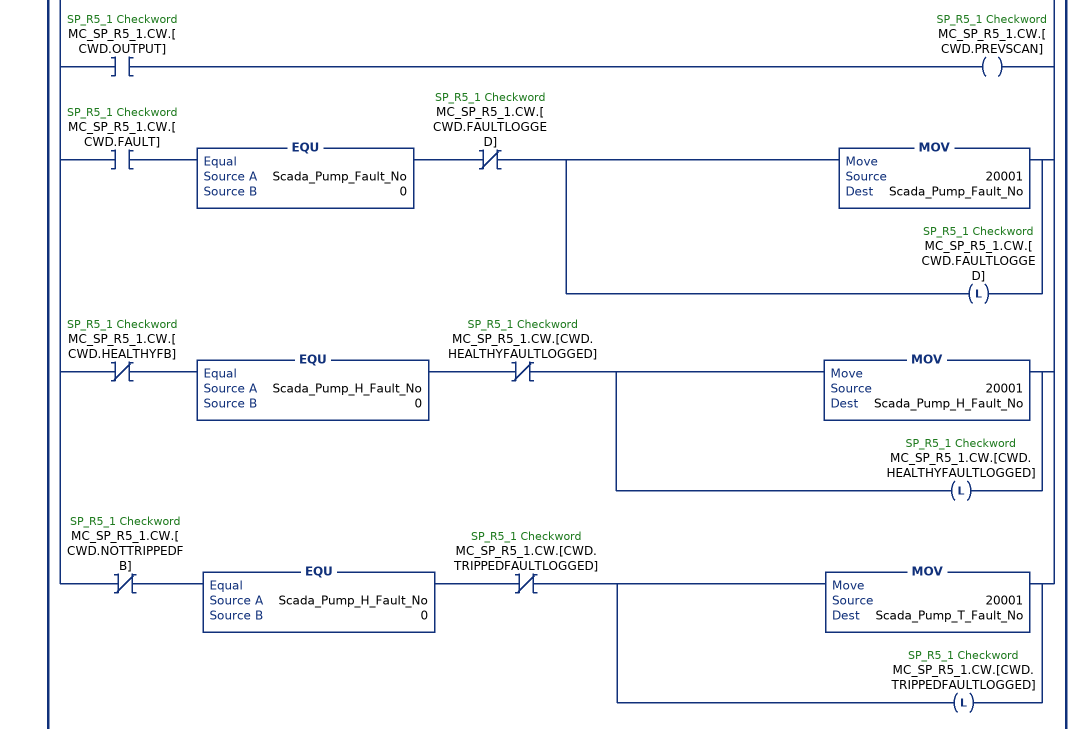
   7: [NEQ(MC_SP_R5_1.DriveBits,0) OTE(MC_SP_R5_1.CW.[CWD.AUTODRV]) ,[XIC(MC_SP_R5_1.CW.[CWD.AUTODRV]) XIO(MC_SP_R5_1.CW.[CWD.MANUAL]) ,XIC(MC_SP_R5_1.CW.[CWD.MANDRV]) XIC(MC_SP_R5_1.CW.[CWD.MANUAL]) ] OTE(MC_SP_R5_1.CW.[CWD.OUTPUT]) ,XIC(MC_SP_R5_1.CW.[CWD.OUTPUT]) OTE(MC_SP_R5_1_D) ,XIC(S:FS) [OTU(MC_SP_R5_1.CW.[CWD.MANUAL]) ,LEQ(MC_SP_R5_1.CheckTime,0) MOV(Default_Check_Time,MC_SP_R5_1.CheckTime) ] ,[[XIC(MC_SP_R5_1_R) XIO(Item_Simulation_Flag) ,XIC(Item_Simulation_Flag) [XIC(MC_SP_R5_1.CW.[CWD.OUTPUT]) XIO(MC_SP_R5_1.CW.[CWD.SIMFAIL]) ,XIO(MC_SP_R5_1.CW.[CWD.OUTPUT]) XIC(MC_SP_R5_1.CW.[CWD.SIMFAIL]) ] ] OTE(MC_SP_R5_1.CW.[CWD.RUNFB]) ,[XIC(Item_Simulation_Flag) ,XIC(MC_SP_R5_1.CW.[CWD.CHECKOFF]) ,XIC(Unused_Healthy_Feedback) ] OTE(MC_SP_R5_1.CW.[CWD.HEALTHYFB]) ,[XIC(Item_Simulation_Flag) ,XIC(MC_SP_R5_1.CW.[CWD.CHECKOFF]) ,XIC(Unused_NotTripped_Feedback) ] OTE(MC_SP_R5_1.CW.[CWD.NOTTRIPPEDFB]) ] ,[XIC(MC_SP_R5_1.CW.[CWD.OUTPUT]) XIO(MC_SP_R5_1.CW.[CWD.PREVSCAN]) ,XIO(MC_SP_R5_1.CW.[CWD.OUTPUT]) XIC(MC_SP_R5_1.CW.[CWD.PREVSCAN]) ] CLR(MC_SP_R5_1.CheckTimer) ,XIC(One_Second_One_Scan) LES(MC_SP_R5_1.CheckTimer,MC_SP_R5_1.CheckTime) ADD(MC_SP_R5_1.CheckTimer,1,MC_SP_R5_1.CheckTimer) ,XIO(MC_SP_R5_1.CW.[CWD.FAULT]) OTU(MC_SP_R5_1.CW.[CWD.FAULTLOGGED]) ,[GEQ(MC_SP_R5_1.CheckTimer,MC_SP_R5_1.CheckTime) [XIC(MC_SP_R5_1.CW.[CWD.OUTPUT]) XIO(MC_SP_R5_1.CW.[CWD.RUNFB]) ,XIO(MC_SP_R5_1.CW.[CWD.OUTPUT]) XIC(MC_SP_R5_1.CW.[CWD.RUNFB]) ] ,XIO(MC_SP_R5_1.CW.[CWD.HEALTHYFB]) ,XIO(MC_SP_R5_1.CW.[CWD.NOTTRIPPEDFB]) ,XIC(MC_SP_R5_1.CW.[CWD.FAULT]) XIC(Item_Faults_Are_Latched) ,XIC(MC_SP_R5_1.CW.[CWD.HIGHLIGHT]) ] XIO(MC_SP_R5_1.CW.[CWD.CHECKOFF]) XIO(Alarm_Reset) [OTE(MC_SP_R5_1.CW.[CWD.FAULT]) ,ALMD(MC_SP_R5_1_ALARM,0,0,0,0) ] ,XIC(MC_SP_R5_1.CW.[CWD.OUTPUT]) OTE(MC_SP_R5_1.CW.[CWD.PREVSCAN]) ,XIC(MC_SP_R5_1.CW.[CWD.FAULT]) EQU(Scada_Pump_Fault_No,0) XIO(MC_SP_R5_1.CW.[CWD.FAULTLOGGED]) [MOV(20001,Scada_Pump_Fault_No) ,OTL(MC_SP_R5_1.CW.[CWD.FAULTLOGGED]) ] ,XIO(MC_SP_R5_1.CW.[CWD.HEALTHYFB]) EQU(Scada_Pump_H_Fault_No,0) XIO(MC_SP_R5_1.CW.[CWD.HEALTHYFAULTLOGGED]) [MOV(20001,Scada_Pump_H_Fault_No) ,OTL(MC_SP_R5_1.CW.[CWD.HEALTHYFAULTLOGGED]) ] ,XIO(MC_SP_R5_1.CW.[CWD.NOTTRIPPEDFB]) EQU(Scada_Pump_H_Fault_No,0) XIO(MC_SP_R5_1.CW.[CWD.TRIPPEDFAULTLOGGED]) [MOV(20001,Scada_Pump_T_Fault_No) ,OTL(MC_SP_R5_1.CW.[CWD.TRIPPEDFAULTLOGGED]) ] ];
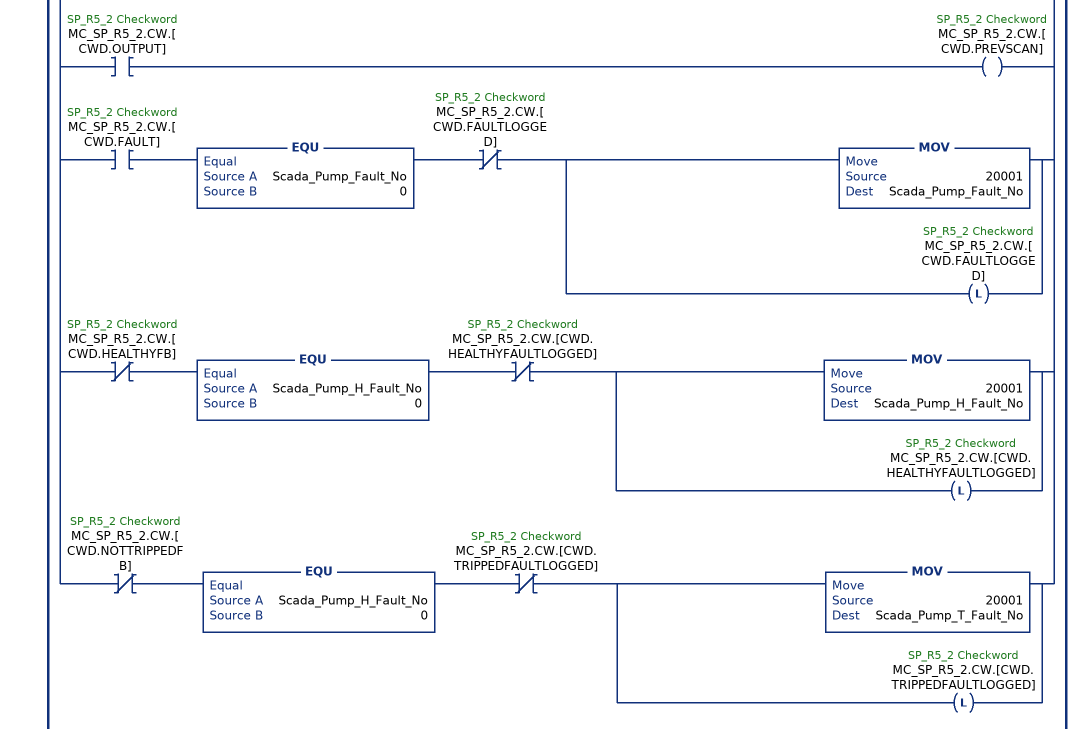
   8: [NEQ(MC_SP_R5_2.DriveBits,0) OTE(MC_SP_R5_2.CW.[CWD.AUTODRV]) ,[XIC(MC_SP_R5_2.CW.[CWD.AUTODRV]) XIO(MC_SP_R5_2.CW.[CWD.MANUAL]) ,XIC(MC_SP_R5_2.CW.[CWD.MANDRV]) XIC(MC_SP_R5_2.CW.[CWD.MANUAL]) ] OTE(MC_SP_R5_2.CW.[CWD.OUTPUT]) ,XIC(MC_SP_R5_2.CW.[CWD.OUTPUT]) OTE(MC_SP_R5_2_D) ,XIC(S:FS) [OTU(MC_SP_R5_2.CW.[CWD.MANUAL]) ,LEQ(MC_SP_R5_2.CheckTime,0) MOV(Default_Check_Time,MC_SP_R5_2.CheckTime) ] ,[[XIC(MC_SP_R5_2_R) XIO(Item_Simulation_Flag) ,XIC(Item_Simulation_Flag) [XIC(MC_SP_R5_2.CW.[CWD.OUTPUT]) XIO(MC_SP_R5_2.CW.[CWD.SIMFAIL]) ,XIO(MC_SP_R5_2.CW.[CWD.OUTPUT]) XIC(MC_SP_R5_2.CW.[CWD.SIMFAIL]) ] ] OTE(MC_SP_R5_2.CW.[CWD.RUNFB]) ,[XIC(Item_Simulation_Flag) ,XIC(MC_SP_R5_2.CW.[CWD.CHECKOFF]) ,XIC(Unused_Healthy_Feedback) ] OTE(MC_SP_R5_2.CW.[CWD.HEALTHYFB]) ,[XIC(Item_Simulation_Flag) ,XIC(MC_SP_R5_2.CW.[CWD.CHECKOFF]) ,XIC(Unused_NotTripped_Feedback) ] OTE(MC_SP_R5_2.CW.[CWD.NOTTRIPPEDFB]) ] ,[XIC(MC_SP_R5_2.CW.[CWD.OUTPUT]) XIO(MC_SP_R5_2.CW.[CWD.PREVSCAN]) ,XIO(MC_SP_R5_2.CW.[CWD.OUTPUT]) XIC(MC_SP_R5_2.CW.[CWD.PREVSCAN]) ] CLR(MC_SP_R5_2.CheckTimer) ,XIC(One_Second_One_Scan) LES(MC_SP_R5_2.CheckTimer,MC_SP_R5_2.CheckTime) ADD(MC_SP_R5_2.CheckTimer,1,MC_SP_R5_2.CheckTimer) ,XIO(MC_SP_R5_2.CW.[CWD.FAULT]) OTU(MC_SP_R5_2.CW.[CWD.FAULTLOGGED]) ,[GEQ(MC_SP_R5_2.CheckTimer,MC_SP_R5_2.CheckTime) [XIC(MC_SP_R5_2.CW.[CWD.OUTPUT]) XIO(MC_SP_R5_2.CW.[CWD.RUNFB]) ,XIO(MC_SP_R5_2.CW.[CWD.OUTPUT]) XIC(MC_SP_R5_2.CW.[CWD.RUNFB]) ] ,XIO(MC_SP_R5_2.CW.[CWD.HEALTHYFB]) ,XIO(MC_SP_R5_2.CW.[CWD.NOTTRIPPEDFB]) ,XIC(MC_SP_R5_2.CW.[CWD.FAULT]) XIC(Item_Faults_Are_Latched) ,XIC(MC_SP_R5_2.CW.[CWD.HIGHLIGHT]) ] XIO(MC_SP_R5_2.CW.[CWD.CHECKOFF]) XIO(Alarm_Reset) [OTE(MC_SP_R5_2.CW.[CWD.FAULT]) ,ALMD(MC_SP_R5_2_ALARM,0,0,0,0) ] ,XIC(MC_SP_R5_2.CW.[CWD.OUTPUT]) OTE(MC_SP_R5_2.CW.[CWD.PREVSCAN]) ,XIC(MC_SP_R5_2.CW.[CWD.FAULT]) EQU(Scada_Pump_Fault_No,0) XIO(MC_SP_R5_2.CW.[CWD.FAULTLOGGED]) [MOV(20001,Scada_Pump_Fault_No) ,OTL(MC_SP_R5_2.CW.[CWD.FAULTLOGGED]) ] ,XIO(MC_SP_R5_2.CW.[CWD.HEALTHYFB]) EQU(Scada_Pump_H_Fault_No,0) XIO(MC_SP_R5_2.CW.[CWD.HEALTHYFAULTLOGGED]) [MOV(20001,Scada_Pump_H_Fault_No) ,OTL(MC_SP_R5_2.CW.[CWD.HEALTHYFAULTLOGGED]) ] ,XIO(MC_SP_R5_2.CW.[CWD.NOTTRIPPEDFB]) EQU(Scada_Pump_H_Fault_No,0) XIO(MC_SP_R5_2.CW.[CWD.TRIPPEDFAULTLOGGED]) [MOV(20001,Scada_Pump_T_Fault_No) ,OTL(MC_SP_R5_2.CW.[CWD.TRIPPEDFAULTLOGGED]) ] ];
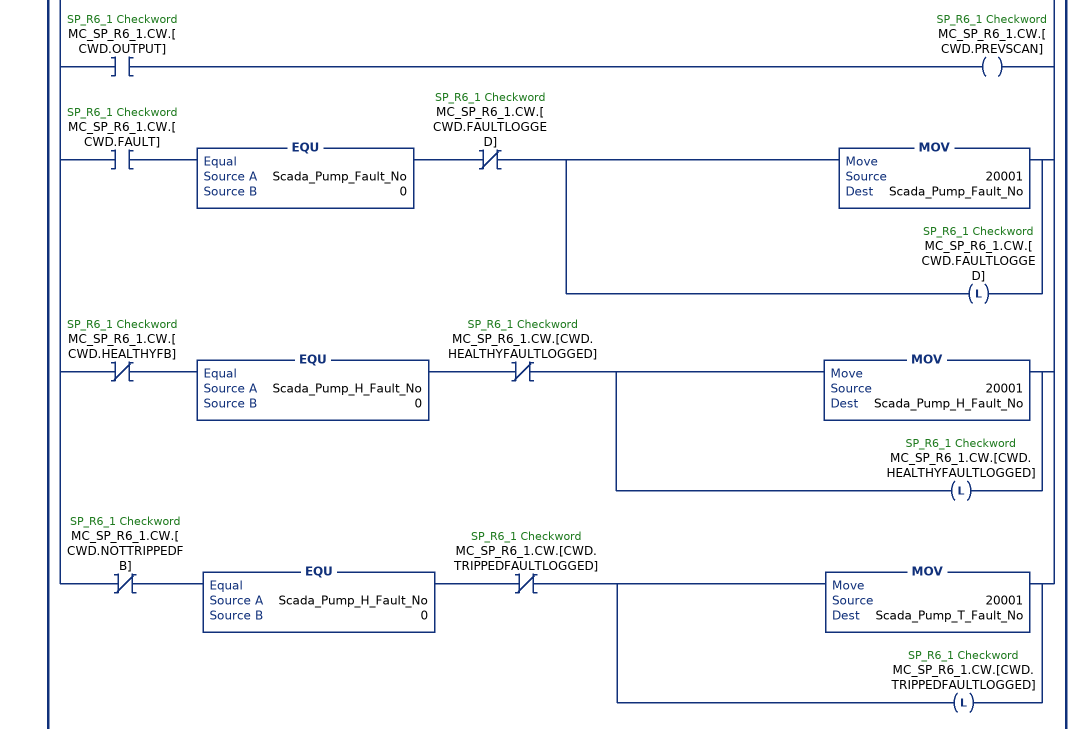
   9: [NEQ(MC_SP_R6_1.DriveBits,0) OTE(MC_SP_R6_1.CW.[CWD.AUTODRV]) ,[XIC(MC_SP_R6_1.CW.[CWD.AUTODRV]) XIO(MC_SP_R6_1.CW.[CWD.MANUAL]) ,XIC(MC_SP_R6_1.CW.[CWD.MANDRV]) XIC(MC_SP_R6_1.CW.[CWD.MANUAL]) ] OTE(MC_SP_R6_1.CW.[CWD.OUTPUT]) ,XIC(MC_SP_R6_1.CW.[CWD.OUTPUT]) OTE(MC_SP_R6_1_D) ,XIC(S:FS) [OTU(MC_SP_R6_1.CW.[CWD.MANUAL]) ,LEQ(MC_SP_R6_1.CheckTime,0) MOV(Default_Check_Time,MC_SP_R6_1.CheckTime) ] ,[[XIC(MC_SP_R6_1_R) XIO(Item_Simulation_Flag) ,XIC(Item_Simulation_Flag) [XIC(MC_SP_R6_1.CW.[CWD.OUTPUT]) XIO(MC_SP_R6_1.CW.[CWD.SIMFAIL]) ,XIO(MC_SP_R6_1.CW.[CWD.OUTPUT]) XIC(MC_SP_R6_1.CW.[CWD.SIMFAIL]) ] ] OTE(MC_SP_R6_1.CW.[CWD.RUNFB]) ,[XIC(Item_Simulation_Flag) ,XIC(MC_SP_R6_1.CW.[CWD.CHECKOFF]) ,XIC(Unused_Healthy_Feedback) ] OTE(MC_SP_R6_1.CW.[CWD.HEALTHYFB]) ,[XIC(Item_Simulation_Flag) ,XIC(MC_SP_R6_1.CW.[CWD.CHECKOFF]) ,XIC(Unused_NotTripped_Feedback) ] OTE(MC_SP_R6_1.CW.[CWD.NOTTRIPPEDFB]) ] ,[XIC(MC_SP_R6_1.CW.[CWD.OUTPUT]) XIO(MC_SP_R6_1.CW.[CWD.PREVSCAN]) ,XIO(MC_SP_R6_1.CW.[CWD.OUTPUT]) XIC(MC_SP_R6_1.CW.[CWD.PREVSCAN]) ] CLR(MC_SP_R6_1.CheckTimer) ,XIC(One_Second_One_Scan) LES(MC_SP_R6_1.CheckTimer,MC_SP_R6_1.CheckTime) ADD(MC_SP_R6_1.CheckTimer,1,MC_SP_R6_1.CheckTimer) ,XIO(MC_SP_R6_1.CW.[CWD.FAULT]) OTU(MC_SP_R6_1.CW.[CWD.FAULTLOGGED]) ,[GEQ(MC_SP_R6_1.CheckTimer,MC_SP_R6_1.CheckTime) [XIC(MC_SP_R6_1.CW.[CWD.OUTPUT]) XIO(MC_SP_R6_1.CW.[CWD.RUNFB]) ,XIO(MC_SP_R6_1.CW.[CWD.OUTPUT]) XIC(MC_SP_R6_1.CW.[CWD.RUNFB]) ] ,XIO(MC_SP_R6_1.CW.[CWD.HEALTHYFB]) ,XIO(MC_SP_R6_1.CW.[CWD.NOTTRIPPEDFB]) ,XIC(MC_SP_R6_1.CW.[CWD.FAULT]) XIC(Item_Faults_Are_Latched) ,XIC(MC_SP_R6_1.CW.[CWD.HIGHLIGHT]) ] XIO(MC_SP_R6_1.CW.[CWD.CHECKOFF]) XIO(Alarm_Reset) [OTE(MC_SP_R6_1.CW.[CWD.FAULT]) ,ALMD(MC_SP_R6_1_ALARM,0,0,0,0) ] ,XIC(MC_SP_R6_1.CW.[CWD.OUTPUT]) OTE(MC_SP_R6_1.CW.[CWD.PREVSCAN]) ,XIC(MC_SP_R6_1.CW.[CWD.FAULT]) EQU(Scada_Pump_Fault_No,0) XIO(MC_SP_R6_1.CW.[CWD.FAULTLOGGED]) [MOV(20001,Scada_Pump_Fault_No) ,OTL(MC_SP_R6_1.CW.[CWD.FAULTLOGGED]) ] ,XIO(MC_SP_R6_1.CW.[CWD.HEALTHYFB]) EQU(Scada_Pump_H_Fault_No,0) XIO(MC_SP_R6_1.CW.[CWD.HEALTHYFAULTLOGGED]) [MOV(20001,Scada_Pump_H_Fault_No) ,OTL(MC_SP_R6_1.CW.[CWD.HEALTHYFAULTLOGGED]) ] ,XIO(MC_SP_R6_1.CW.[CWD.NOTTRIPPEDFB]) EQU(Scada_Pump_H_Fault_No,0) XIO(MC_SP_R6_1.CW.[CWD.TRIPPEDFAULTLOGGED]) [MOV(20001,Scada_Pump_T_Fault_No) ,OTL(MC_SP_R6_1.CW.[CWD.TRIPPEDFAULTLOGGED]) ] ];
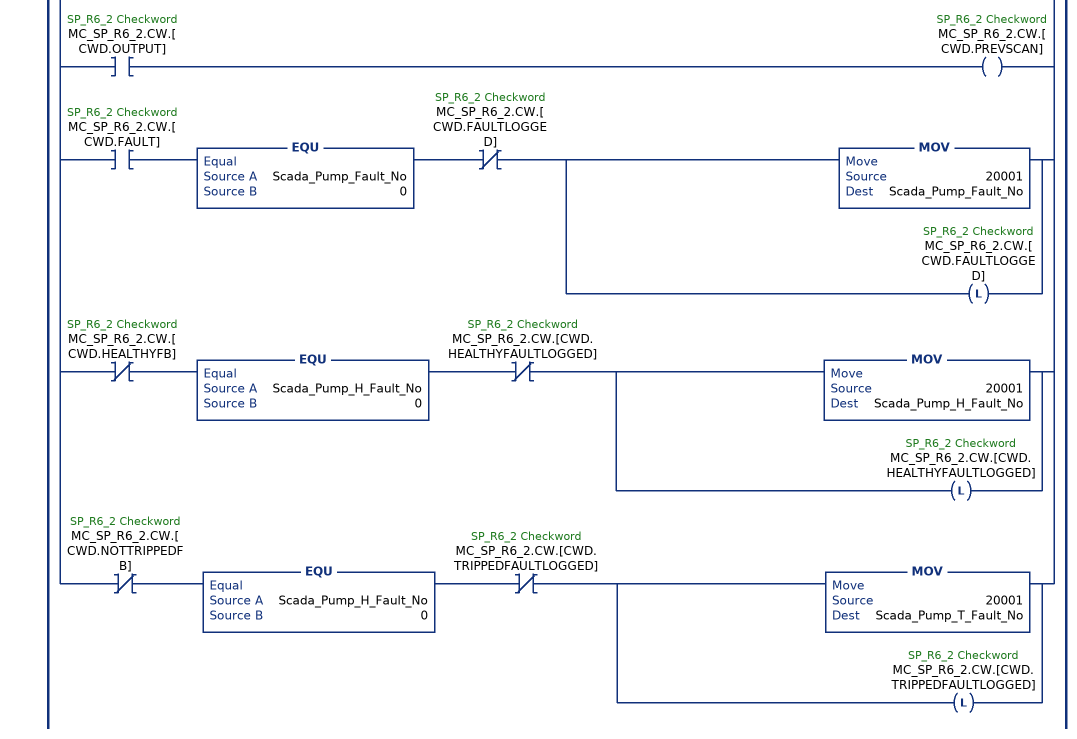
   10: [NEQ(MC_SP_R6_2.DriveBits,0) OTE(MC_SP_R6_2.CW.[CWD.AUTODRV]) ,[XIC(MC_SP_R6_2.CW.[CWD.AUTODRV]) XIO(MC_SP_R6_2.CW.[CWD.MANUAL]) ,XIC(MC_SP_R6_2.CW.[CWD.MANDRV]) XIC(MC_SP_R6_2.CW.[CWD.MANUAL]) ] OTE(MC_SP_R6_2.CW.[CWD.OUTPUT]) ,XIC(MC_SP_R6_2.CW.[CWD.OUTPUT]) OTE(MC_SP_R6_2_D) ,XIC(S:FS) [OTU(MC_SP_R6_2.CW.[CWD.MANUAL]) ,LEQ(MC_SP_R6_2.CheckTime,0) MOV(Default_Check_Time,MC_SP_R6_2.CheckTime) ] ,[[XIC(MC_SP_R6_2_R) XIO(Item_Simulation_Flag) ,XIC(Item_Simulation_Flag) [XIC(MC_SP_R6_2.CW.[CWD.OUTPUT]) XIO(MC_SP_R6_2.CW.[CWD.SIMFAIL]) ,XIO(MC_SP_R6_2.CW.[CWD.OUTPUT]) XIC(MC_SP_R6_2.CW.[CWD.SIMFAIL]) ] ] OTE(MC_SP_R6_2.CW.[CWD.RUNFB]) ,[XIC(Item_Simulation_Flag) ,XIC(MC_SP_R6_2.CW.[CWD.CHECKOFF]) ,XIC(Unused_Healthy_Feedback) ] OTE(MC_SP_R6_2.CW.[CWD.HEALTHYFB]) ,[XIC(Item_Simulation_Flag) ,XIC(MC_SP_R6_2.CW.[CWD.CHECKOFF]) ,XIC(Unused_NotTripped_Feedback) ] OTE(MC_SP_R6_2.CW.[CWD.NOTTRIPPEDFB]) ] ,[XIC(MC_SP_R6_2.CW.[CWD.OUTPUT]) XIO(MC_SP_R6_2.CW.[CWD.PREVSCAN]) ,XIO(MC_SP_R6_2.CW.[CWD.OUTPUT]) XIC(MC_SP_R6_2.CW.[CWD.PREVSCAN]) ] CLR(MC_SP_R6_2.CheckTimer) ,XIC(One_Second_One_Scan) LES(MC_SP_R6_2.CheckTimer,MC_SP_R6_2.CheckTime) ADD(MC_SP_R6_2.CheckTimer,1,MC_SP_R6_2.CheckTimer) ,XIO(MC_SP_R6_2.CW.[CWD.FAULT]) OTU(MC_SP_R6_2.CW.[CWD.FAULTLOGGED]) ,[GEQ(MC_SP_R6_2.CheckTimer,MC_SP_R6_2.CheckTime) [XIC(MC_SP_R6_2.CW.[CWD.OUTPUT]) XIO(MC_SP_R6_2.CW.[CWD.RUNFB]) ,XIO(MC_SP_R6_2.CW.[CWD.OUTPUT]) XIC(MC_SP_R6_2.CW.[CWD.RUNFB]) ] ,XIO(MC_SP_R6_2.CW.[CWD.HEALTHYFB]) ,XIO(MC_SP_R6_2.CW.[CWD.NOTTRIPPEDFB]) ,XIC(MC_SP_R6_2.CW.[CWD.FAULT]) XIC(Item_Faults_Are_Latched) ,XIC(MC_SP_R6_2.CW.[CWD.HIGHLIGHT]) ] XIO(MC_SP_R6_2.CW.[CWD.CHECKOFF]) XIO(Alarm_Reset) [OTE(MC_SP_R6_2.CW.[CWD.FAULT]) ,ALMD(MC_SP_R6_2_ALARM,0,0,0,0) ] ,XIC(MC_SP_R6_2.CW.[CWD.OUTPUT]) OTE(MC_SP_R6_2.CW.[CWD.PREVSCAN]) ,XIC(MC_SP_R6_2.CW.[CWD.FAULT]) EQU(Scada_Pump_Fault_No,0) XIO(MC_SP_R6_2.CW.[CWD.FAULTLOGGED]) [MOV(20001,Scada_Pump_Fault_No) ,OTL(MC_SP_R6_2.CW.[CWD.FAULTLOGGED]) ] ,XIO(MC_SP_R6_2.CW.[CWD.HEALTHYFB]) EQU(Scada_Pump_H_Fault_No,0) XIO(MC_SP_R6_2.CW.[CWD.HEALTHYFAULTLOGGED]) [MOV(20001,Scada_Pump_H_Fault_No) ,OTL(MC_SP_R6_2.CW.[CWD.HEALTHYFAULTLOGGED]) ] ,XIO(MC_SP_R6_2.CW.[CWD.NOTTRIPPEDFB]) EQU(Scada_Pump_H_Fault_No,0) XIO(MC_SP_R6_2.CW.[CWD.TRIPPEDFAULTLOGGED]) [MOV(20001,Scada_Pump_T_Fault_No) ,OTL(MC_SP_R6_2.CW.[CWD.TRIPPEDFAULTLOGGED]) ] ];
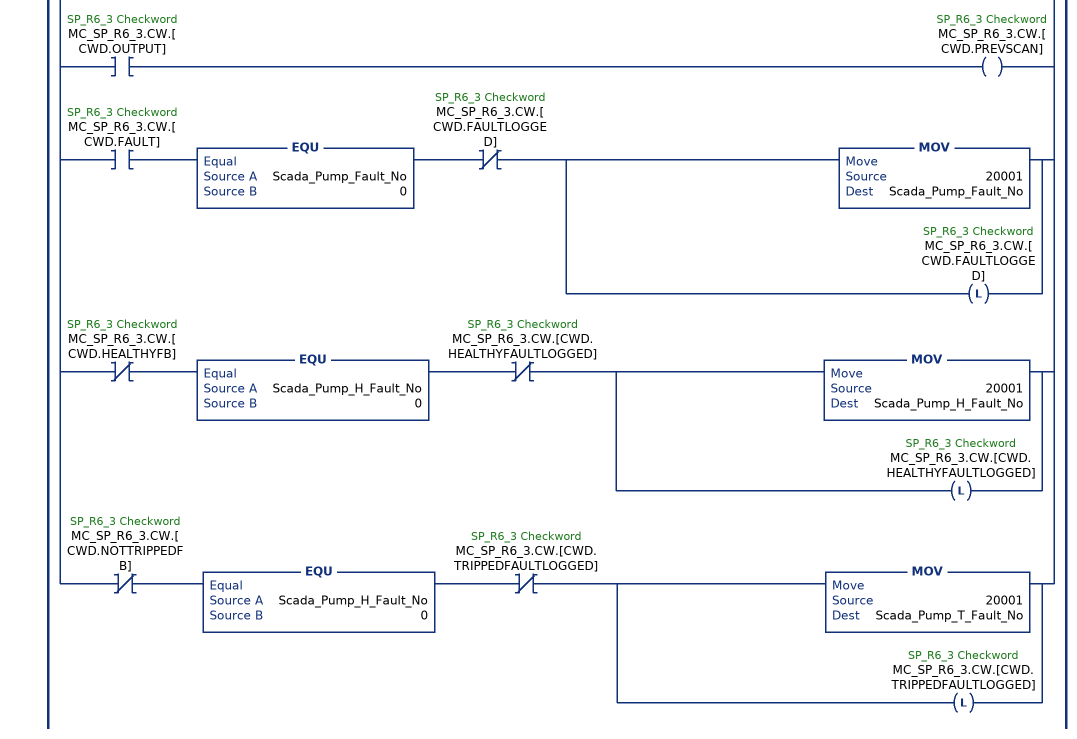
   11: [NEQ(MC_SP_R6_3.DriveBits,0) OTE(MC_SP_R6_3.CW.[CWD.AUTODRV]) ,[XIC(MC_SP_R6_3.CW.[CWD.AUTODRV]) XIO(MC_SP_R6_3.CW.[CWD.MANUAL]) ,XIC(MC_SP_R6_3.CW.[CWD.MANDRV]) XIC(MC_SP_R6_3.CW.[CWD.MANUAL]) ] OTE(MC_SP_R6_3.CW.[CWD.OUTPUT]) ,XIC(MC_SP_R6_3.CW.[CWD.OUTPUT]) OTE(MC_SP_R6_3_D) ,XIC(S:FS) [OTU(MC_SP_R6_3.CW.[CWD.MANUAL]) ,LEQ(MC_SP_R6_3.CheckTime,0) MOV(Default_Check_Time,MC_SP_R6_3.CheckTime) ] ,[[XIC(MC_SP_R6_3_R) XIO(Item_Simulation_Flag) ,XIC(Item_Simulation_Flag) [XIC(MC_SP_R6_3.CW.[CWD.OUTPUT]) XIO(MC_SP_R6_3.CW.[CWD.SIMFAIL]) ,XIO(MC_SP_R6_3.CW.[CWD.OUTPUT]) XIC(MC_SP_R6_3.CW.[CWD.SIMFAIL]) ] ] OTE(MC_SP_R6_3.CW.[CWD.RUNFB]) ,[XIC(Item_Simulation_Flag) ,XIC(MC_SP_R6_3.CW.[CWD.CHECKOFF]) ,XIC(Unused_Healthy_Feedback) ] OTE(MC_SP_R6_3.CW.[CWD.HEALTHYFB]) ,[XIC(Item_Simulation_Flag) ,XIC(MC_SP_R6_3.CW.[CWD.CHECKOFF]) ,XIC(Unused_NotTripped_Feedback) ] OTE(MC_SP_R6_3.CW.[CWD.NOTTRIPPEDFB]) ] ,[XIC(MC_SP_R6_3.CW.[CWD.OUTPUT]) XIO(MC_SP_R6_3.CW.[CWD.PREVSCAN]) ,XIO(MC_SP_R6_3.CW.[CWD.OUTPUT]) XIC(MC_SP_R6_3.CW.[CWD.PREVSCAN]) ] CLR(MC_SP_R6_3.CheckTimer) ,XIC(One_Second_One_Scan) LES(MC_SP_R6_3.CheckTimer,MC_SP_R6_3.CheckTime) ADD(MC_SP_R6_3.CheckTimer,1,MC_SP_R6_3.CheckTimer) ,XIO(MC_SP_R6_3.CW.[CWD.FAULT]) OTU(MC_SP_R6_3.CW.[CWD.FAULTLOGGED]) ,[GEQ(MC_SP_R6_3.CheckTimer,MC_SP_R6_3.CheckTime) [XIC(MC_SP_R6_3.CW.[CWD.OUTPUT]) XIO(MC_SP_R6_3.CW.[CWD.RUNFB]) ,XIO(MC_SP_R6_3.CW.[CWD.OUTPUT]) XIC(MC_SP_R6_3.CW.[CWD.RUNFB]) ] ,XIO(MC_SP_R6_3.CW.[CWD.HEALTHYFB]) ,XIO(MC_SP_R6_3.CW.[CWD.NOTTRIPPEDFB]) ,XIC(MC_SP_R6_3.CW.[CWD.FAULT]) XIC(Item_Faults_Are_Latched) ,XIC(MC_SP_R6_3.CW.[CWD.HIGHLIGHT]) ] XIO(MC_SP_R6_3.CW.[CWD.CHECKOFF]) XIO(Alarm_Reset) [OTE(MC_SP_R6_3.CW.[CWD.FAULT]) ,ALMD(MC_SP_R6_3_ALARM,0,0,0,0) ] ,XIC(MC_SP_R6_3.CW.[CWD.OUTPUT]) OTE(MC_SP_R6_3.CW.[CWD.PREVSCAN]) ,XIC(MC_SP_R6_3.CW.[CWD.FAULT]) EQU(Scada_Pump_Fault_No,0) XIO(MC_SP_R6_3.CW.[CWD.FAULTLOGGED]) [MOV(20001,Scada_Pump_Fault_No) ,OTL(MC_SP_R6_3.CW.[CWD.FAULTLOGGED]) ] ,XIO(MC_SP_R6_3.CW.[CWD.HEALTHYFB]) EQU(Scada_Pump_H_Fault_No,0) XIO(MC_SP_R6_3.CW.[CWD.HEALTHYFAULTLOGGED]) [MOV(20001,Scada_Pump_H_Fault_No) ,OTL(MC_SP_R6_3.CW.[CWD.HEALTHYFAULTLOGGED]) ] ,XIO(MC_SP_R6_3.CW.[CWD.NOTTRIPPEDFB]) EQU(Scada_Pump_H_Fault_No,0) XIO(MC_SP_R6_3.CW.[CWD.TRIPPEDFAULTLOGGED]) [MOV(20001,Scada_Pump_T_Fault_No) ,OTL(MC_SP_R6_3.CW.[CWD.TRIPPEDFAULTLOGGED]) ] ];
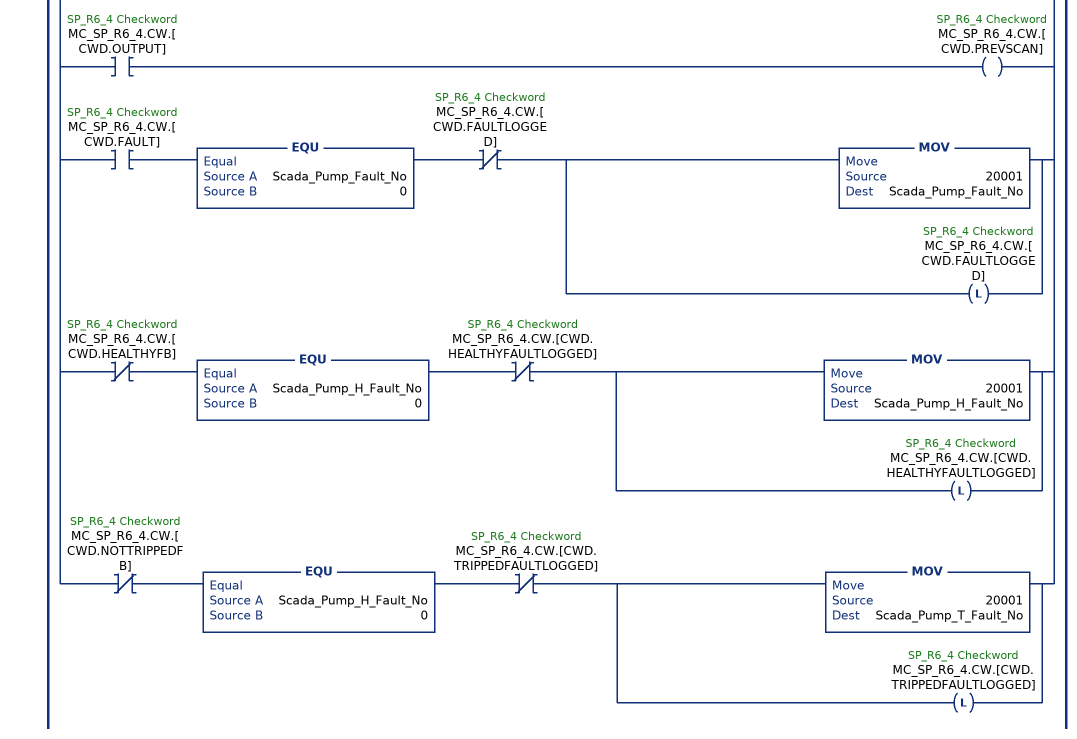
   12: [NEQ(MC_SP_R6_4.DriveBits,0) OTE(MC_SP_R6_4.CW.[CWD.AUTODRV]) ,[XIC(MC_SP_R6_4.CW.[CWD.AUTODRV]) XIO(MC_SP_R6_4.CW.[CWD.MANUAL]) ,XIC(MC_SP_R6_4.CW.[CWD.MANDRV]) XIC(MC_SP_R6_4.CW.[CWD.MANUAL]) ] OTE(MC_SP_R6_4.CW.[CWD.OUTPUT]) ,XIC(MC_SP_R6_4.CW.[CWD.OUTPUT]) OTE(MC_SP_R6_4_D) ,XIC(S:FS) [OTU(MC_SP_R6_4.CW.[CWD.MANUAL]) ,LEQ(MC_SP_R6_4.CheckTime,0) MOV(Default_Check_Time,MC_SP_R6_4.CheckTime) ] ,[[XIC(MC_SP_R6_4_R) XIO(Item_Simulation_Flag) ,XIC(Item_Simulation_Flag) [XIC(MC_SP_R6_4.CW.[CWD.OUTPUT]) XIO(MC_SP_R6_4.CW.[CWD.SIMFAIL]) ,XIO(MC_SP_R6_4.CW.[CWD.OUTPUT]) XIC(MC_SP_R6_4.CW.[CWD.SIMFAIL]) ] ] OTE(MC_SP_R6_4.CW.[CWD.RUNFB]) ,[XIC(Item_Simulation_Flag) ,XIC(MC_SP_R6_4.CW.[CWD.CHECKOFF]) ,XIC(Unused_Healthy_Feedback) ] OTE(MC_SP_R6_4.CW.[CWD.HEALTHYFB]) ,[XIC(Item_Simulation_Flag) ,XIC(MC_SP_R6_4.CW.[CWD.CHECKOFF]) ,XIC(Unused_NotTripped_Feedback) ] OTE(MC_SP_R6_4.CW.[CWD.NOTTRIPPEDFB]) ] ,[XIC(MC_SP_R6_4.CW.[CWD.OUTPUT]) XIO(MC_SP_R6_4.CW.[CWD.PREVSCAN]) ,XIO(MC_SP_R6_4.CW.[CWD.OUTPUT]) XIC(MC_SP_R6_4.CW.[CWD.PREVSCAN]) ] CLR(MC_SP_R6_4.CheckTimer) ,XIC(One_Second_One_Scan) LES(MC_SP_R6_4.CheckTimer,MC_SP_R6_4.CheckTime) ADD(MC_SP_R6_4.CheckTimer,1,MC_SP_R6_4.CheckTimer) ,XIO(MC_SP_R6_4.CW.[CWD.FAULT]) OTU(MC_SP_R6_4.CW.[CWD.FAULTLOGGED]) ,[GEQ(MC_SP_R6_4.CheckTimer,MC_SP_R6_4.CheckTime) [XIC(MC_SP_R6_4.CW.[CWD.OUTPUT]) XIO(MC_SP_R6_4.CW.[CWD.RUNFB]) ,XIO(MC_SP_R6_4.CW.[CWD.OUTPUT]) XIC(MC_SP_R6_4.CW.[CWD.RUNFB]) ] ,XIO(MC_SP_R6_4.CW.[CWD.HEALTHYFB]) ,XIO(MC_SP_R6_4.CW.[CWD.NOTTRIPPEDFB]) ,XIC(MC_SP_R6_4.CW.[CWD.FAULT]) XIC(Item_Faults_Are_Latched) ,XIC(MC_SP_R6_4.CW.[CWD.HIGHLIGHT]) ] XIO(MC_SP_R6_4.CW.[CWD.CHECKOFF]) XIO(Alarm_Reset) [OTE(MC_SP_R6_4.CW.[CWD.FAULT]) ,ALMD(MC_SP_R6_4_ALARM,0,0,0,0) ] ,XIC(MC_SP_R6_4.CW.[CWD.OUTPUT]) OTE(MC_SP_R6_4.CW.[CWD.PREVSCAN]) ,XIC(MC_SP_R6_4.CW.[CWD.FAULT]) EQU(Scada_Pump_Fault_No,0) XIO(MC_SP_R6_4.CW.[CWD.FAULTLOGGED]) [MOV(20001,Scada_Pump_Fault_No) ,OTL(MC_SP_R6_4.CW.[CWD.FAULTLOGGED]) ] ,XIO(MC_SP_R6_4.CW.[CWD.HEALTHYFB]) EQU(Scada_Pump_H_Fault_No,0) XIO(MC_SP_R6_4.CW.[CWD.HEALTHYFAULTLOGGED]) [MOV(20001,Scada_Pump_H_Fault_No) ,OTL(MC_SP_R6_4.CW.[CWD.HEALTHYFAULTLOGGED]) ] ,XIO(MC_SP_R6_4.CW.[CWD.NOTTRIPPEDFB]) EQU(Scada_Pump_H_Fault_No,0) XIO(MC_SP_R6_4.CW.[CWD.TRIPPEDFAULTLOGGED]) [MOV(20001,Scada_Pump_T_Fault_No) ,OTL(MC_SP_R6_4.CW.[CWD.TRIPPEDFAULTLOGGED]) ] ];
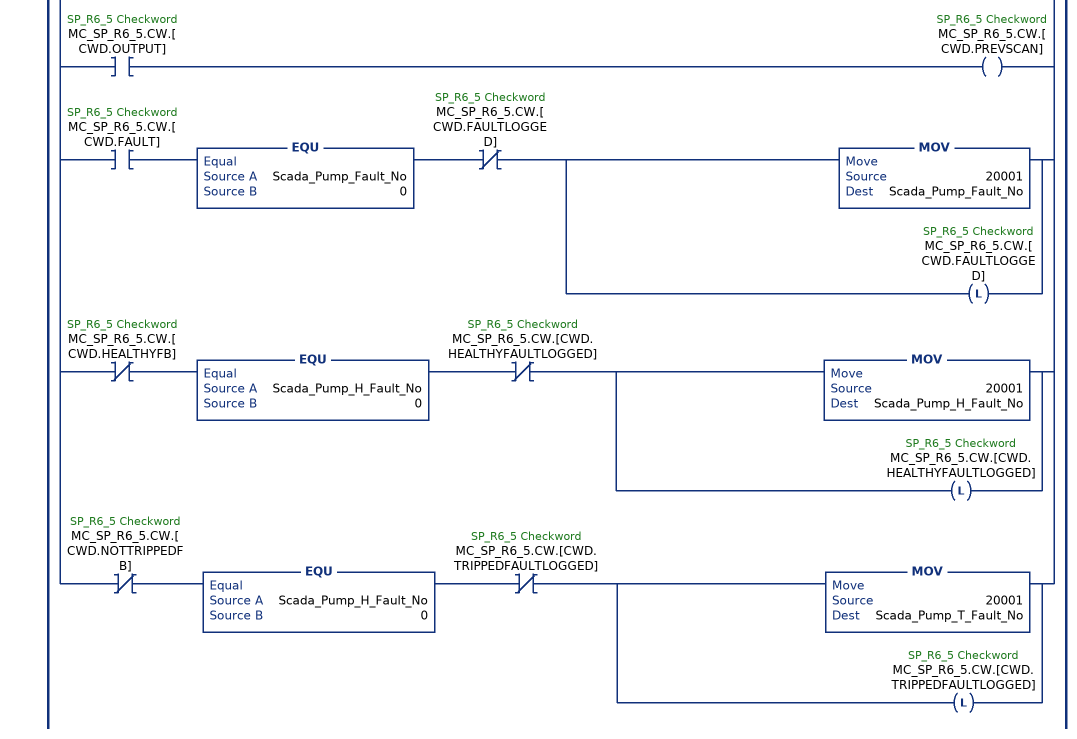
   13: [NEQ(MC_SP_R6_5.DriveBits,0) OTE(MC_SP_R6_5.CW.[CWD.AUTODRV]) ,[XIC(MC_SP_R6_5.CW.[CWD.AUTODRV]) XIO(MC_SP_R6_5.CW.[CWD.MANUAL]) ,XIC(MC_SP_R6_5.CW.[CWD.MANDRV]) XIC(MC_SP_R6_5.CW.[CWD.MANUAL]) ] OTE(MC_SP_R6_5.CW.[CWD.OUTPUT]) ,XIC(MC_SP_R6_5.CW.[CWD.OUTPUT]) OTE(MC_SP_R6_5_D) ,XIC(S:FS) [OTU(MC_SP_R6_5.CW.[CWD.MANUAL]) ,LEQ(MC_SP_R6_5.CheckTime,0) MOV(Default_Check_Time,MC_SP_R6_5.CheckTime) ] ,[[XIC(MC_SP_R6_5_R) XIO(Item_Simulation_Flag) ,XIC(Item_Simulation_Flag) [XIC(MC_SP_R6_5.CW.[CWD.OUTPUT]) XIO(MC_SP_R6_5.CW.[CWD.SIMFAIL]) ,XIO(MC_SP_R6_5.CW.[CWD.OUTPUT]) XIC(MC_SP_R6_5.CW.[CWD.SIMFAIL]) ] ] OTE(MC_SP_R6_5.CW.[CWD.RUNFB]) ,[XIC(Item_Simulation_Flag) ,XIC(MC_SP_R6_5.CW.[CWD.CHECKOFF]) ,XIC(Unused_Healthy_Feedback) ] OTE(MC_SP_R6_5.CW.[CWD.HEALTHYFB]) ,[XIC(Item_Simulation_Flag) ,XIC(MC_SP_R6_5.CW.[CWD.CHECKOFF]) ,XIC(Unused_NotTripped_Feedback) ] OTE(MC_SP_R6_5.CW.[CWD.NOTTRIPPEDFB]) ] ,[XIC(MC_SP_R6_5.CW.[CWD.OUTPUT]) XIO(MC_SP_R6_5.CW.[CWD.PREVSCAN]) ,XIO(MC_SP_R6_5.CW.[CWD.OUTPUT]) XIC(MC_SP_R6_5.CW.[CWD.PREVSCAN]) ] CLR(MC_SP_R6_5.CheckTimer) ,XIC(One_Second_One_Scan) LES(MC_SP_R6_5.CheckTimer,MC_SP_R6_5.CheckTime) ADD(MC_SP_R6_5.CheckTimer,1,MC_SP_R6_5.CheckTimer) ,XIO(MC_SP_R6_5.CW.[CWD.FAULT]) OTU(MC_SP_R6_5.CW.[CWD.FAULTLOGGED]) ,[GEQ(MC_SP_R6_5.CheckTimer,MC_SP_R6_5.CheckTime) [XIC(MC_SP_R6_5.CW.[CWD.OUTPUT]) XIO(MC_SP_R6_5.CW.[CWD.RUNFB]) ,XIO(MC_SP_R6_5.CW.[CWD.OUTPUT]) XIC(MC_SP_R6_5.CW.[CWD.RUNFB]) ] ,XIO(MC_SP_R6_5.CW.[CWD.HEALTHYFB]) ,XIO(MC_SP_R6_5.CW.[CWD.NOTTRIPPEDFB]) ,XIC(MC_SP_R6_5.CW.[CWD.FAULT]) XIC(Item_Faults_Are_Latched) ,XIC(MC_SP_R6_5.CW.[CWD.HIGHLIGHT]) ] XIO(MC_SP_R6_5.CW.[CWD.CHECKOFF]) XIO(Alarm_Reset) [OTE(MC_SP_R6_5.CW.[CWD.FAULT]) ,ALMD(MC_SP_R6_5_ALARM,0,0,0,0) ] ,XIC(MC_SP_R6_5.CW.[CWD.OUTPUT]) OTE(MC_SP_R6_5.CW.[CWD.PREVSCAN]) ,XIC(MC_SP_R6_5.CW.[CWD.FAULT]) EQU(Scada_Pump_Fault_No,0) XIO(MC_SP_R6_5.CW.[CWD.FAULTLOGGED]) [MOV(20001,Scada_Pump_Fault_No) ,OTL(MC_SP_R6_5.CW.[CWD.FAULTLOGGED]) ] ,XIO(MC_SP_R6_5.CW.[CWD.HEALTHYFB]) EQU(Scada_Pump_H_Fault_No,0) XIO(MC_SP_R6_5.CW.[CWD.HEALTHYFAULTLOGGED]) [MOV(20001,Scada_Pump_H_Fault_No) ,OTL(MC_SP_R6_5.CW.[CWD.HEALTHYFAULTLOGGED]) ] ,XIO(MC_SP_R6_5.CW.[CWD.NOTTRIPPEDFB]) EQU(Scada_Pump_H_Fault_No,0) XIO(MC_SP_R6_5.CW.[CWD.TRIPPEDFAULTLOGGED]) [MOV(20001,Scada_Pump_T_Fault_No) ,OTL(MC_SP_R6_5.CW.[CWD.TRIPPEDFAULTLOGGED]) ] ];
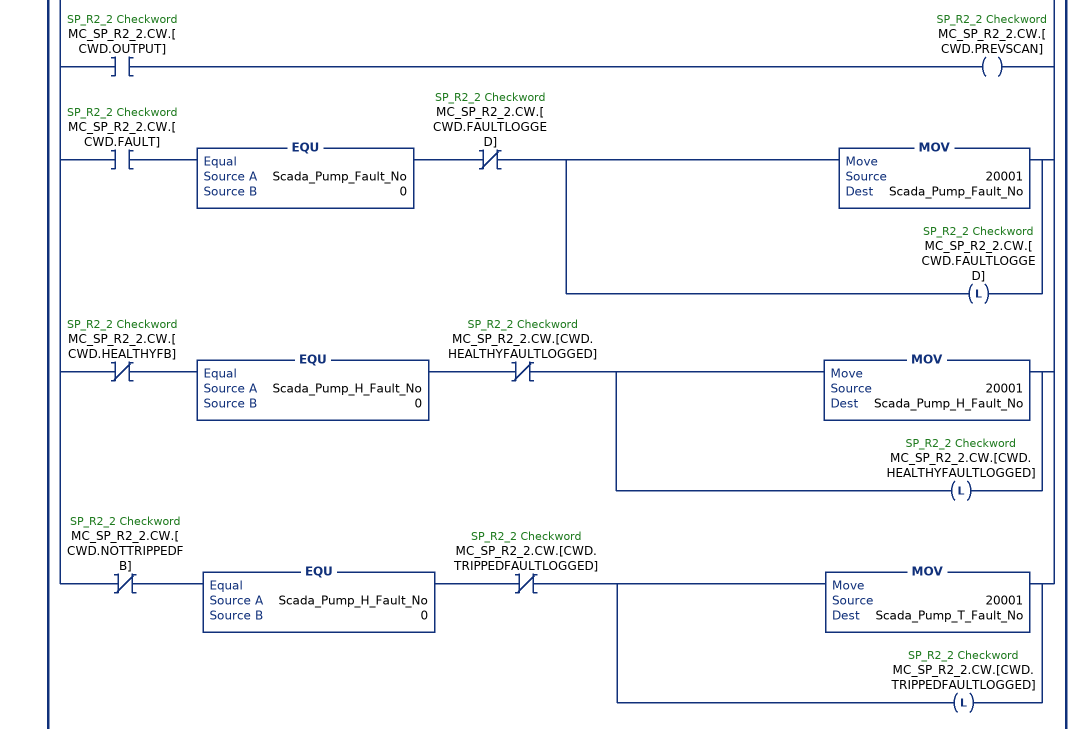
   14: [NEQ(MC_SP_R2_2.DriveBits,0) OTE(MC_SP_R2_2.CW.[CWD.AUTODRV]) ,[XIC(MC_SP_R2_2.CW.[CWD.AUTODRV]) XIO(MC_SP_R2_2.CW.[CWD.MANUAL]) ,XIC(MC_SP_R2_2.CW.[CWD.MANDRV]) XIC(MC_SP_R2_2.CW.[CWD.MANUAL]) ] OTE(MC_SP_R2_2.CW.[CWD.OUTPUT]) ,XIC(MC_SP_R2_2.CW.[CWD.OUTPUT]) OTE(MC_SP_R2_2_D) ,XIC(S:FS) [OTU(MC_SP_R2_2.CW.[CWD.MANUAL]) ,LEQ(MC_SP_R2_2.CheckTime,0) MOV(Default_Check_Time,MC_SP_R2_2.CheckTime) ] ,[[XIC(MC_SP_R2_2_R) XIO(Item_Simulation_Flag) ,XIC(Item_Simulation_Flag) [XIC(MC_SP_R2_2.CW.[CWD.OUTPUT]) XIO(MC_SP_R2_2.CW.[CWD.SIMFAIL]) ,XIO(MC_SP_R2_2.CW.[CWD.OUTPUT]) XIC(MC_SP_R2_2.CW.[CWD.SIMFAIL]) ] ] OTE(MC_SP_R2_2.CW.[CWD.RUNFB]) ,[XIC(Item_Simulation_Flag) ,XIC(MC_SP_R2_2.CW.[CWD.CHECKOFF]) ,XIC(Unused_Healthy_Feedback) ] OTE(MC_SP_R2_2.CW.[CWD.HEALTHYFB]) ,[XIC(Item_Simulation_Flag) ,XIC(MC_SP_R2_2.CW.[CWD.CHECKOFF]) ,XIC(Unused_NotTripped_Feedback) ] OTE(MC_SP_R2_2.CW.[CWD.NOTTRIPPEDFB]) ] ,[XIC(MC_SP_R2_2.CW.[CWD.OUTPUT]) XIO(MC_SP_R2_2.CW.[CWD.PREVSCAN]) ,XIO(MC_SP_R2_2.CW.[CWD.OUTPUT]) XIC(MC_SP_R2_2.CW.[CWD.PREVSCAN]) ] CLR(MC_SP_R2_2.CheckTimer) ,XIC(One_Second_One_Scan) LES(MC_SP_R2_2.CheckTimer,MC_SP_R2_2.CheckTime) ADD(MC_SP_R2_2.CheckTimer,1,MC_SP_R2_2.CheckTimer) ,XIO(MC_SP_R2_2.CW.[CWD.FAULT]) OTU(MC_SP_R2_2.CW.[CWD.FAULTLOGGED]) ,[GEQ(MC_SP_R2_2.CheckTimer,MC_SP_R2_2.CheckTime) [XIC(MC_SP_R2_2.CW.[CWD.OUTPUT]) XIO(MC_SP_R2_2.CW.[CWD.RUNFB]) ,XIO(MC_SP_R2_2.CW.[CWD.OUTPUT]) XIC(MC_SP_R2_2.CW.[CWD.RUNFB]) ] ,XIO(MC_SP_R2_2.CW.[CWD.HEALTHYFB]) ,XIO(MC_SP_R2_2.CW.[CWD.NOTTRIPPEDFB]) ,XIC(MC_SP_R2_2.CW.[CWD.FAULT]) XIC(Item_Faults_Are_Latched) ,XIC(MC_SP_R2_2.CW.[CWD.HIGHLIGHT]) ] XIO(MC_SP_R2_2.CW.[CWD.CHECKOFF]) XIO(Alarm_Reset) [OTE(MC_SP_R2_2.CW.[CWD.FAULT]) ,ALMD(MC_SP_R2_2_ALARM,0,0,0,0) ] ,XIC(MC_SP_R2_2.CW.[CWD.OUTPUT]) OTE(MC_SP_R2_2.CW.[CWD.PREVSCAN]) ,XIC(MC_SP_R2_2.CW.[CWD.FAULT]) EQU(Scada_Pump_Fault_No,0) XIO(MC_SP_R2_2.CW.[CWD.FAULTLOGGED]) [MOV(20001,Scada_Pump_Fault_No) ,OTL(MC_SP_R2_2.CW.[CWD.FAULTLOGGED]) ] ,XIO(MC_SP_R2_2.CW.[CWD.HEALTHYFB]) EQU(Scada_Pump_H_Fault_No,0) XIO(MC_SP_R2_2.CW.[CWD.HEALTHYFAULTLOGGED]) [MOV(20001,Scada_Pump_H_Fault_No) ,OTL(MC_SP_R2_2.CW.[CWD.HEALTHYFAULTLOGGED]) ] ,XIO(MC_SP_R2_2.CW.[CWD.NOTTRIPPEDFB]) EQU(Scada_Pump_H_Fault_No,0) XIO(MC_SP_R2_2.CW.[CWD.TRIPPEDFAULTLOGGED]) [MOV(20001,Scada_Pump_T_Fault_No) ,OTL(MC_SP_R2_2.CW.[CWD.TRIPPEDFAULTLOGGED]) ] ];
END_ROUTINE
